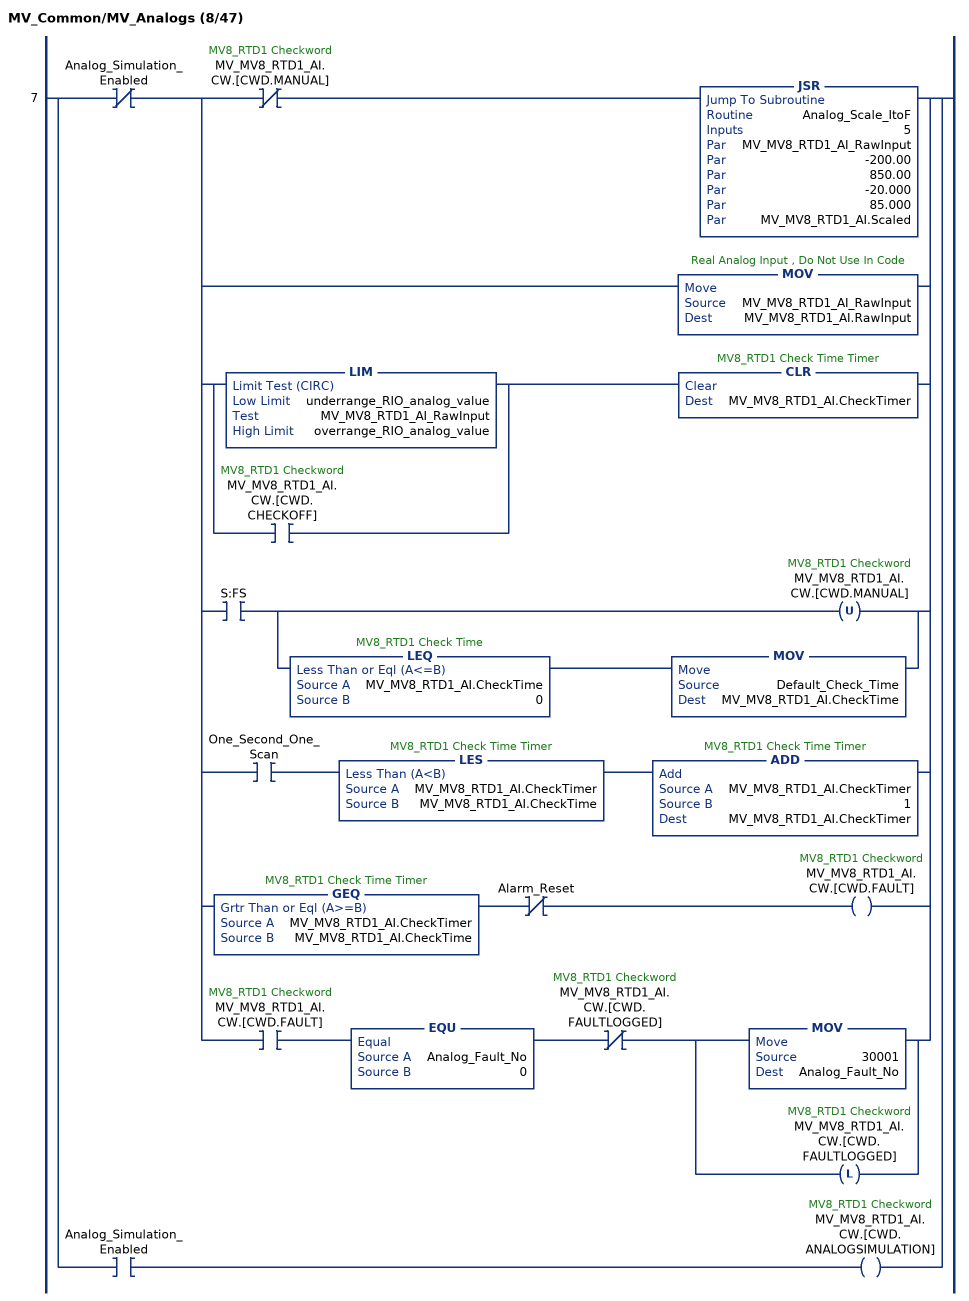
   7: [XIO(Analog_Simulation_Enabled) [XIO(MV_MV8_RTD1_AI.CW.[CWD.MANUAL]) JSR(Analog_Scale_ItoF,5,MV_MV8_RTD1_AI_RawInput,-200.00,850.00,-20.000,85.000,MV_MV8_RTD1_AI.Scaled) ,MOV(MV_MV8_RTD1_AI_RawInput,MV_MV8_RTD1_AI.RawInput) ,[LIM(underrange_RIO_analog_value,MV_MV8_RTD1_AI_RawInput,overrange_RIO_analog_value) ,XIC(MV_MV8_RTD1_AI.CW.[CWD.CHECKOFF]) ] CLR(MV_MV8_RTD1_AI.CheckTimer) ,XIC(S:FS) [OTU(MV_MV8_RTD1_AI.CW.[CWD.MANUAL]) ,LEQ(MV_MV8_RTD1_AI.CheckTime,0) MOV(Default_Check_Time,MV_MV8_RTD1_AI.CheckTime) ] ,XIC(One_Second_One_Scan) LES(MV_MV8_RTD1_AI.CheckTimer,MV_MV8_RTD1_AI.CheckTime) ADD(MV_MV8_RTD1_AI.CheckTimer,1,MV_MV8_RTD1_AI.CheckTimer) ,GEQ(MV_MV8_RTD1_AI.CheckTimer,MV_MV8_RTD1_AI.CheckTime) XIO(Alarm_Reset) OTE(MV_MV8_RTD1_AI.CW.[CWD.FAULT]) ,XIC(MV_MV8_RTD1_AI.CW.[CWD.FAULT]) EQU(Analog_Fault_No,0) XIO(MV_MV8_RTD1_AI.CW.[CWD.FAULTLOGGED]) [MOV(30001,Analog_Fault_No) ,OTL(MV_MV8_RTD1_AI.CW.[CWD.FAULTLOGGED]) ] ] ,XIC(Analog_Simulation_Enabled) OTE(MV_MV8_RTD1_AI.CW.[CWD.ANALOGSIMULATION]) ];
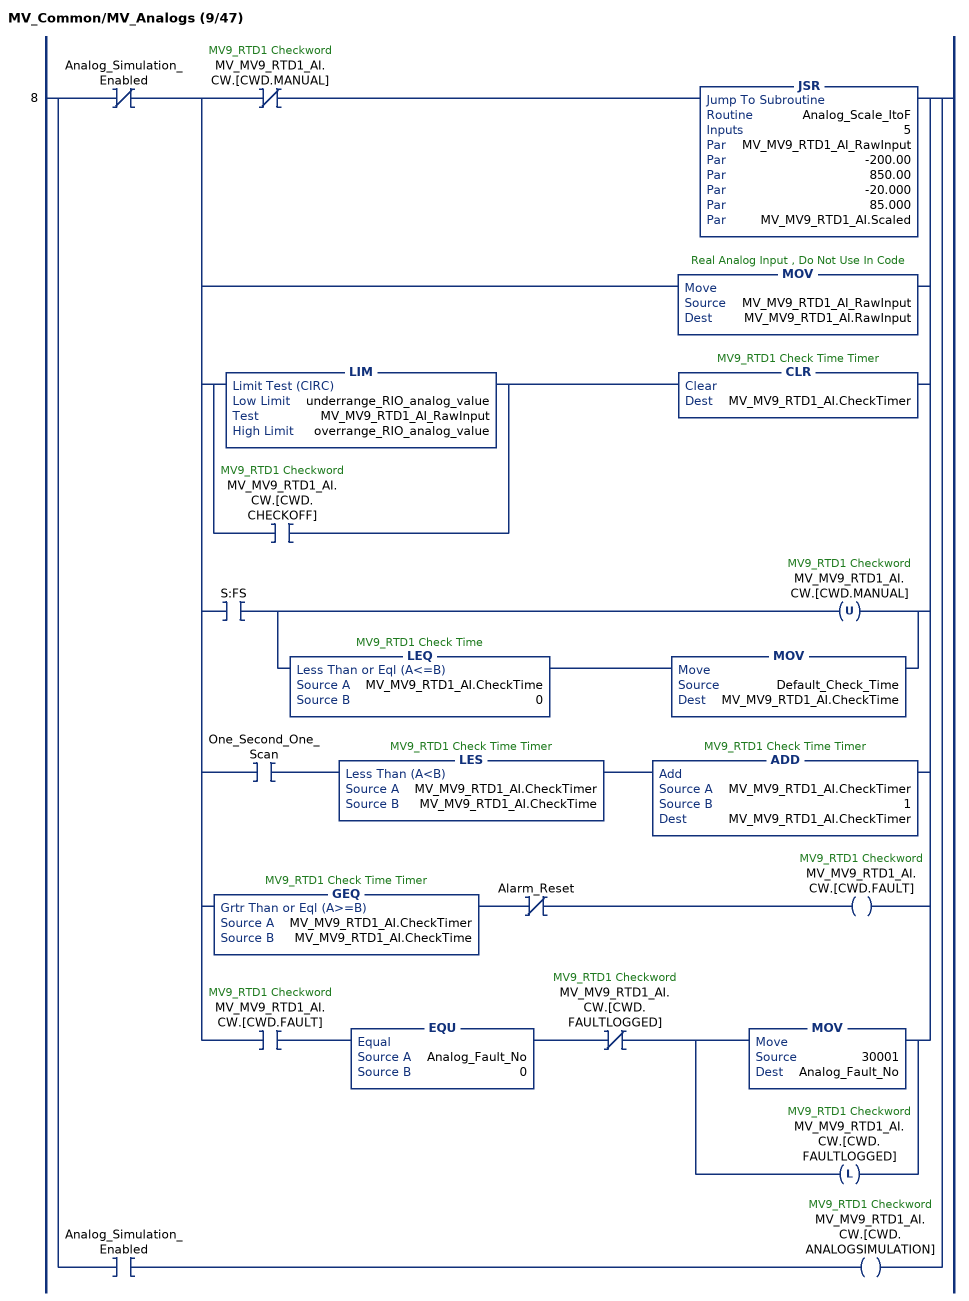
   8: [XIO(Analog_Simulation_Enabled) [XIO(MV_MV9_RTD1_AI.CW.[CWD.MANUAL]) JSR(Analog_Scale_ItoF,5,MV_MV9_RTD1_AI_RawInput,-200.00,850.00,-20.000,85.000,MV_MV9_RTD1_AI.Scaled) ,MOV(MV_MV9_RTD1_AI_RawInput,MV_MV9_RTD1_AI.RawInput) ,[LIM(underrange_RIO_analog_value,MV_MV9_RTD1_AI_RawInput,overrange_RIO_analog_value) ,XIC(MV_MV9_RTD1_AI.CW.[CWD.CHECKOFF]) ] CLR(MV_MV9_RTD1_AI.CheckTimer) ,XIC(S:FS) [OTU(MV_MV9_RTD1_AI.CW.[CWD.MANUAL]) ,LEQ(MV_MV9_RTD1_AI.CheckTime,0) MOV(Default_Check_Time,MV_MV9_RTD1_AI.CheckTime) ] ,XIC(One_Second_One_Scan) LES(MV_MV9_RTD1_AI.CheckTimer,MV_MV9_RTD1_AI.CheckTime) ADD(MV_MV9_RTD1_AI.CheckTimer,1,MV_MV9_RTD1_AI.CheckTimer) ,GEQ(MV_MV9_RTD1_AI.CheckTimer,MV_MV9_RTD1_AI.CheckTime) XIO(Alarm_Reset) OTE(MV_MV9_RTD1_AI.CW.[CWD.FAULT]) ,XIC(MV_MV9_RTD1_AI.CW.[CWD.FAULT]) EQU(Analog_Fault_No,0) XIO(MV_MV9_RTD1_AI.CW.[CWD.FAULTLOGGED]) [MOV(30001,Analog_Fault_No) ,OTL(MV_MV9_RTD1_AI.CW.[CWD.FAULTLOGGED]) ] ] ,XIC(Analog_Simulation_Enabled) OTE(MV_MV9_RTD1_AI.CW.[CWD.ANALOGSIMULATION]) ];
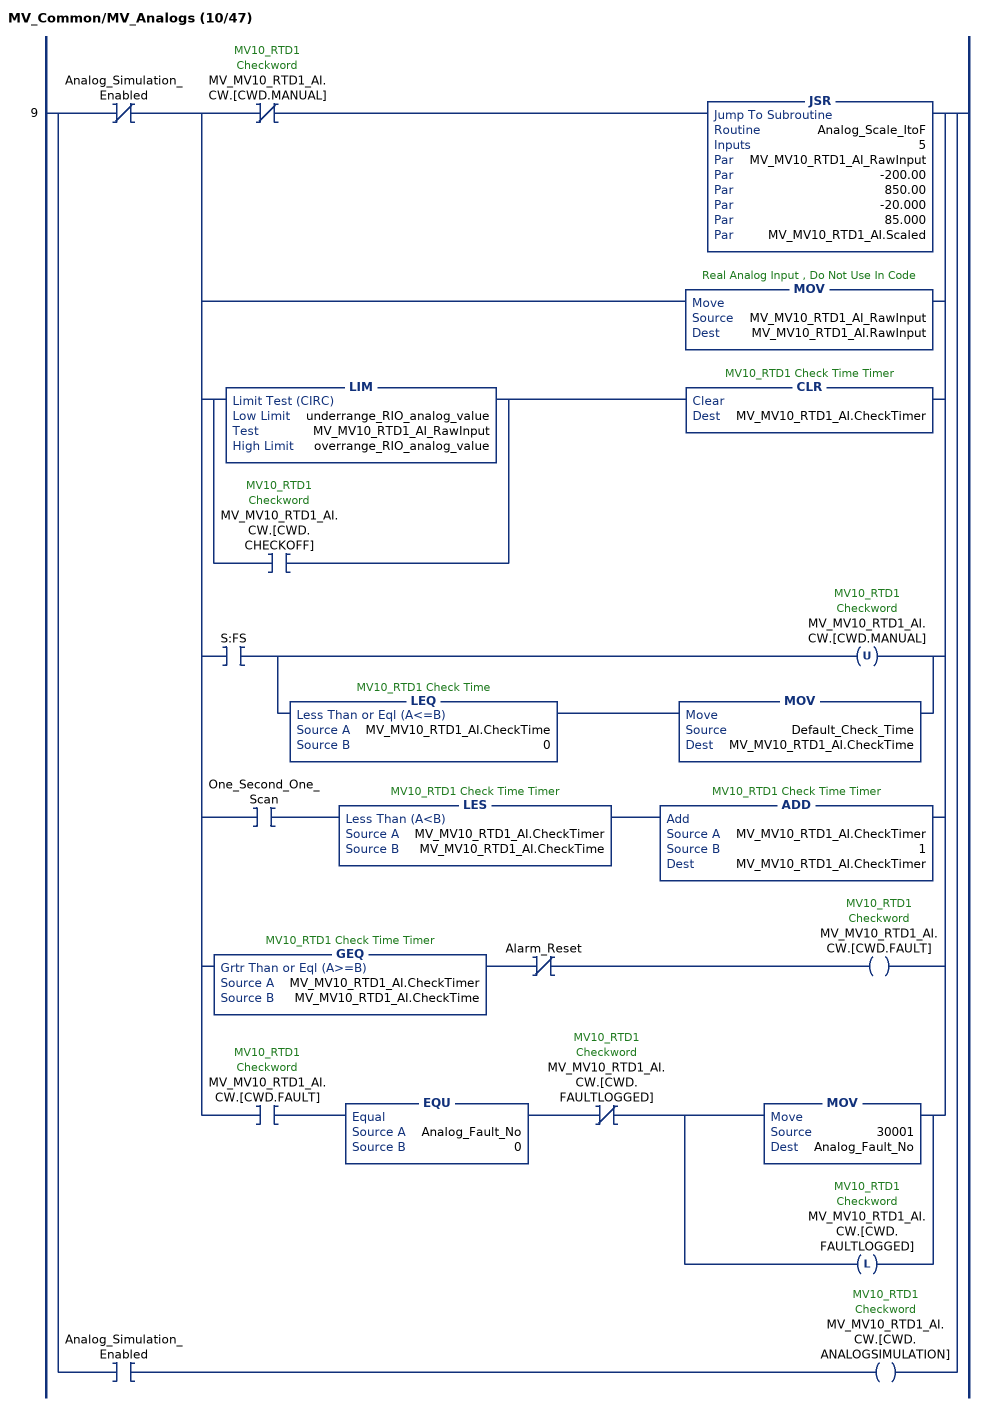
   9: [XIO(Analog_Simulation_Enabled) [XIO(MV_MV10_RTD1_AI.CW.[CWD.MANUAL]) JSR(Analog_Scale_ItoF,5,MV_MV10_RTD1_AI_RawInput,-200.00,850.00,-20.000,85.000,MV_MV10_RTD1_AI.Scaled) ,MOV(MV_MV10_RTD1_AI_RawInput,MV_MV10_RTD1_AI.RawInput) ,[LIM(underrange_RIO_analog_value,MV_MV10_RTD1_AI_RawInput,overrange_RIO_analog_value) ,XIC(MV_MV10_RTD1_AI.CW.[CWD.CHECKOFF]) ] CLR(MV_MV10_RTD1_AI.CheckTimer) ,XIC(S:FS) [OTU(MV_MV10_RTD1_AI.CW.[CWD.MANUAL]) ,LEQ(MV_MV10_RTD1_AI.CheckTime,0) MOV(Default_Check_Time,MV_MV10_RTD1_AI.CheckTime) ] ,XIC(One_Second_One_Scan) LES(MV_MV10_RTD1_AI.CheckTimer,MV_MV10_RTD1_AI.CheckTime) ADD(MV_MV10_RTD1_AI.CheckTimer,1,MV_MV10_RTD1_AI.CheckTimer) ,GEQ(MV_MV10_RTD1_AI.CheckTimer,MV_MV10_RTD1_AI.CheckTime) XIO(Alarm_Reset) OTE(MV_MV10_RTD1_AI.CW.[CWD.FAULT]) ,XIC(MV_MV10_RTD1_AI.CW.[CWD.FAULT]) EQU(Analog_Fault_No,0) XIO(MV_MV10_RTD1_AI.CW.[CWD.FAULTLOGGED]) [MOV(30001,Analog_Fault_No) ,OTL(MV_MV10_RTD1_AI.CW.[CWD.FAULTLOGGED]) ] ] ,XIC(Analog_Simulation_Enabled) OTE(MV_MV10_RTD1_AI.CW.[CWD.ANALOGSIMULATION]) ];
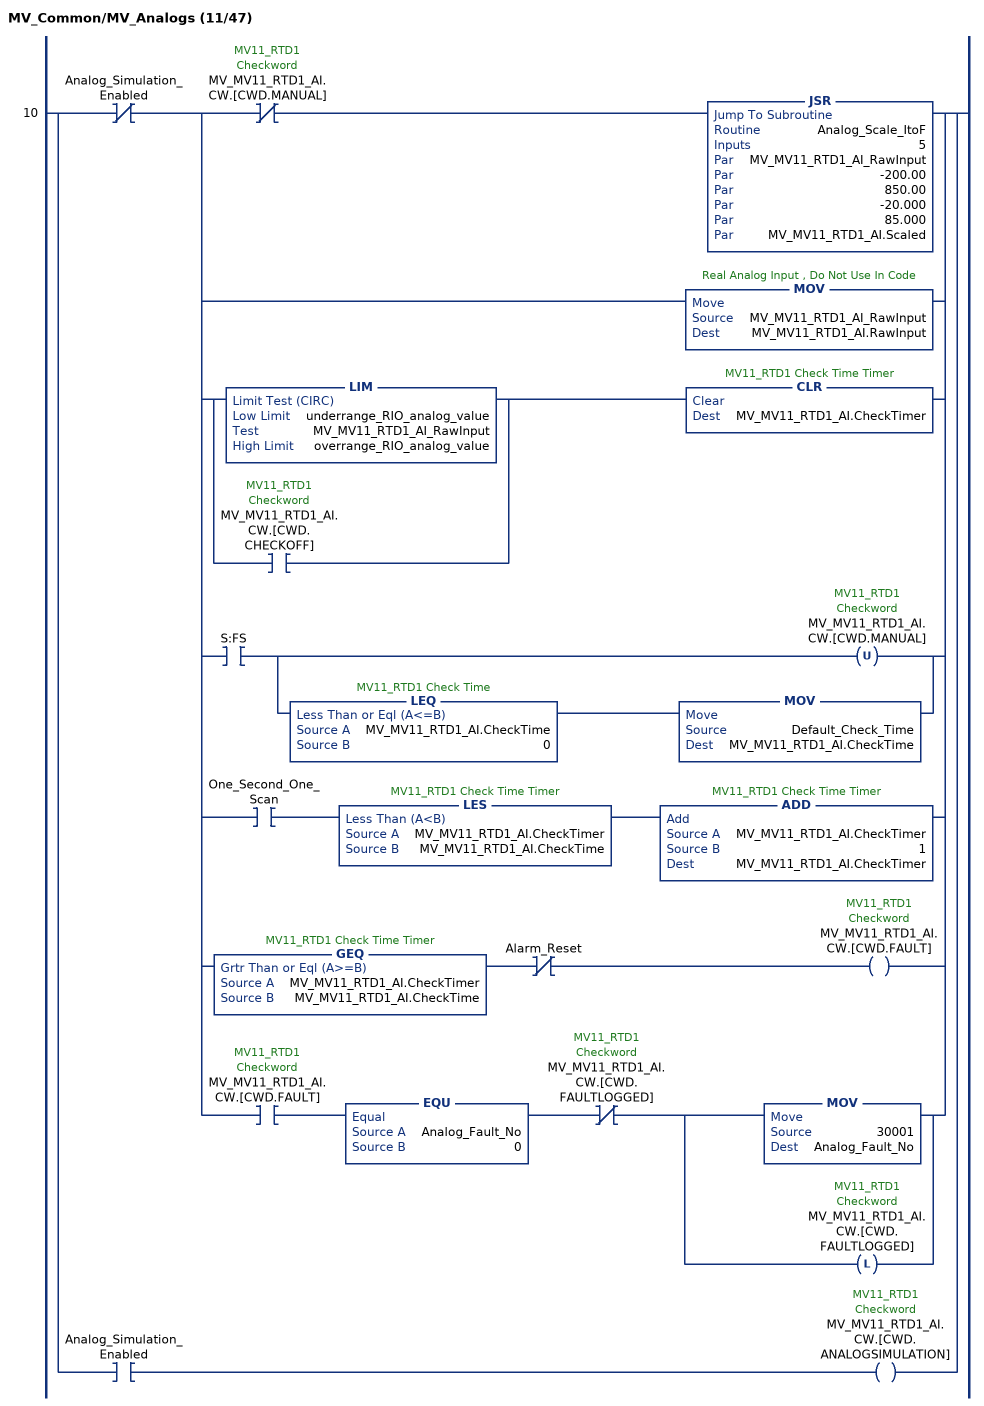
   10: [XIO(Analog_Simulation_Enabled) [XIO(MV_MV11_RTD1_AI.CW.[CWD.MANUAL]) JSR(Analog_Scale_ItoF,5,MV_MV11_RTD1_AI_RawInput,-200.00,850.00,-20.000,85.000,MV_MV11_RTD1_AI.Scaled) ,MOV(MV_MV11_RTD1_AI_RawInput,MV_MV11_RTD1_AI.RawInput) ,[LIM(underrange_RIO_analog_value,MV_MV11_RTD1_AI_RawInput,overrange_RIO_analog_value) ,XIC(MV_MV11_RTD1_AI.CW.[CWD.CHECKOFF]) ] CLR(MV_MV11_RTD1_AI.CheckTimer) ,XIC(S:FS) [OTU(MV_MV11_RTD1_AI.CW.[CWD.MANUAL]) ,LEQ(MV_MV11_RTD1_AI.CheckTime,0) MOV(Default_Check_Time,MV_MV11_RTD1_AI.CheckTime) ] ,XIC(One_Second_One_Scan) LES(MV_MV11_RTD1_AI.CheckTimer,MV_MV11_RTD1_AI.CheckTime) ADD(MV_MV11_RTD1_AI.CheckTimer,1,MV_MV11_RTD1_AI.CheckTimer) ,GEQ(MV_MV11_RTD1_AI.CheckTimer,MV_MV11_RTD1_AI.CheckTime) XIO(Alarm_Reset) OTE(MV_MV11_RTD1_AI.CW.[CWD.FAULT]) ,XIC(MV_MV11_RTD1_AI.CW.[CWD.FAULT]) EQU(Analog_Fault_No,0) XIO(MV_MV11_RTD1_AI.CW.[CWD.FAULTLOGGED]) [MOV(30001,Analog_Fault_No) ,OTL(MV_MV11_RTD1_AI.CW.[CWD.FAULTLOGGED]) ] ] ,XIC(Analog_Simulation_Enabled) OTE(MV_MV11_RTD1_AI.CW.[CWD.ANALOGSIMULATION]) ];
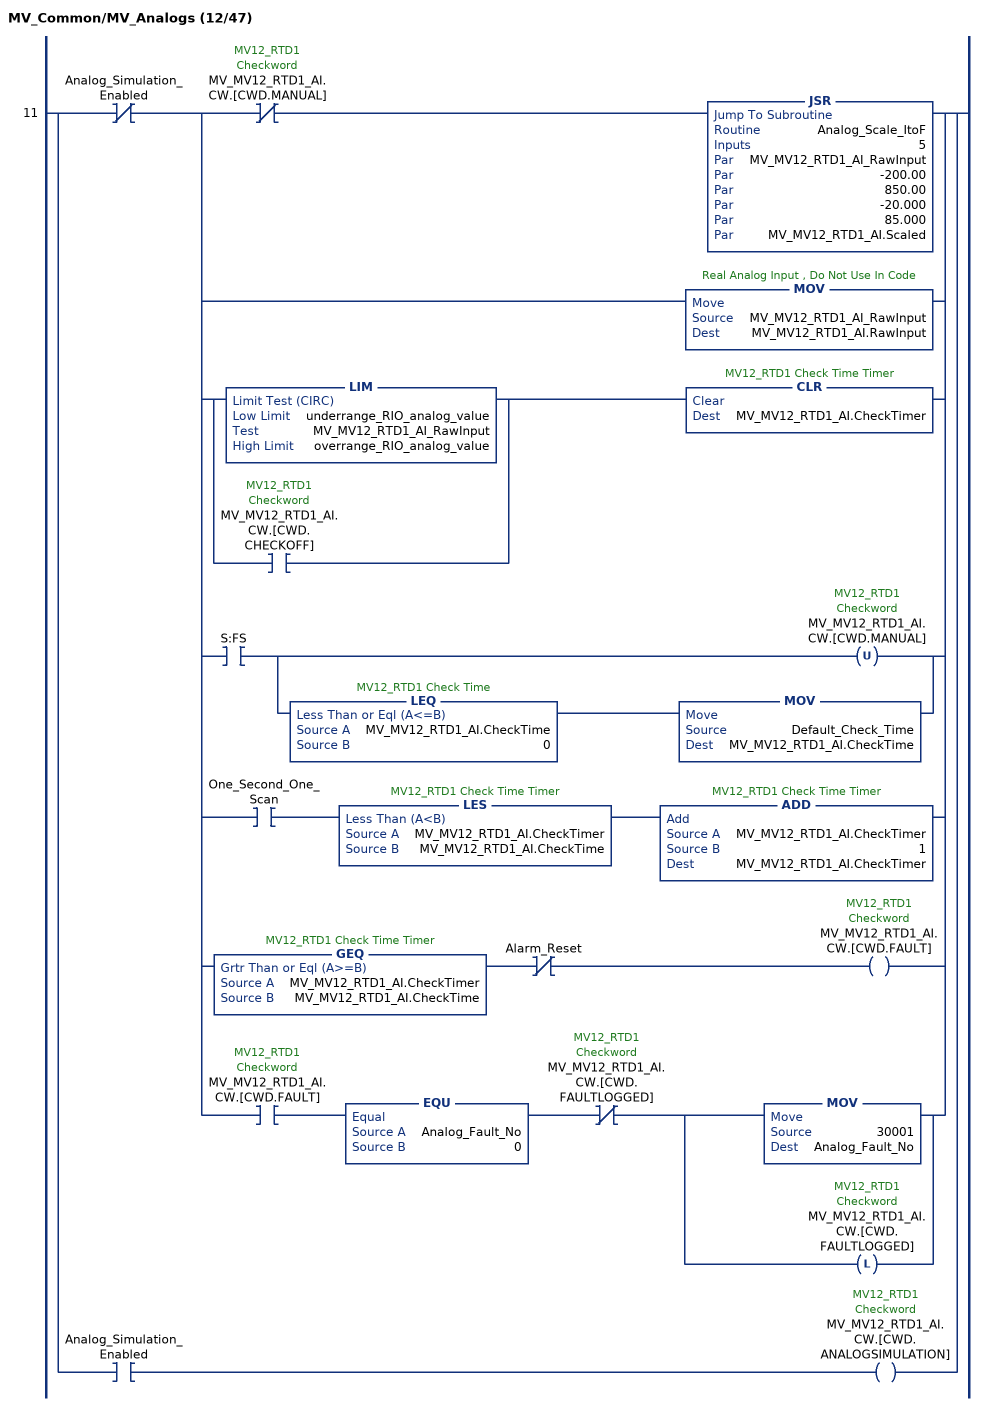
   11: [XIO(Analog_Simulation_Enabled) [XIO(MV_MV12_RTD1_AI.CW.[CWD.MANUAL]) JSR(Analog_Scale_ItoF,5,MV_MV12_RTD1_AI_RawInput,-200.00,850.00,-20.000,85.000,MV_MV12_RTD1_AI.Scaled) ,MOV(MV_MV12_RTD1_AI_RawInput,MV_MV12_RTD1_AI.RawInput) ,[LIM(underrange_RIO_analog_value,MV_MV12_RTD1_AI_RawInput,overrange_RIO_analog_value) ,XIC(MV_MV12_RTD1_AI.CW.[CWD.CHECKOFF]) ] CLR(MV_MV12_RTD1_AI.CheckTimer) ,XIC(S:FS) [OTU(MV_MV12_RTD1_AI.CW.[CWD.MANUAL]) ,LEQ(MV_MV12_RTD1_AI.CheckTime,0) MOV(Default_Check_Time,MV_MV12_RTD1_AI.CheckTime) ] ,XIC(One_Second_One_Scan) LES(MV_MV12_RTD1_AI.CheckTimer,MV_MV12_RTD1_AI.CheckTime) ADD(MV_MV12_RTD1_AI.CheckTimer,1,MV_MV12_RTD1_AI.CheckTimer) ,GEQ(MV_MV12_RTD1_AI.CheckTimer,MV_MV12_RTD1_AI.CheckTime) XIO(Alarm_Reset) OTE(MV_MV12_RTD1_AI.CW.[CWD.FAULT]) ,XIC(MV_MV12_RTD1_AI.CW.[CWD.FAULT]) EQU(Analog_Fault_No,0) XIO(MV_MV12_RTD1_AI.CW.[CWD.FAULTLOGGED]) [MOV(30001,Analog_Fault_No) ,OTL(MV_MV12_RTD1_AI.CW.[CWD.FAULTLOGGED]) ] ] ,XIC(Analog_Simulation_Enabled) OTE(MV_MV12_RTD1_AI.CW.[CWD.ANALOGSIMULATION]) ];
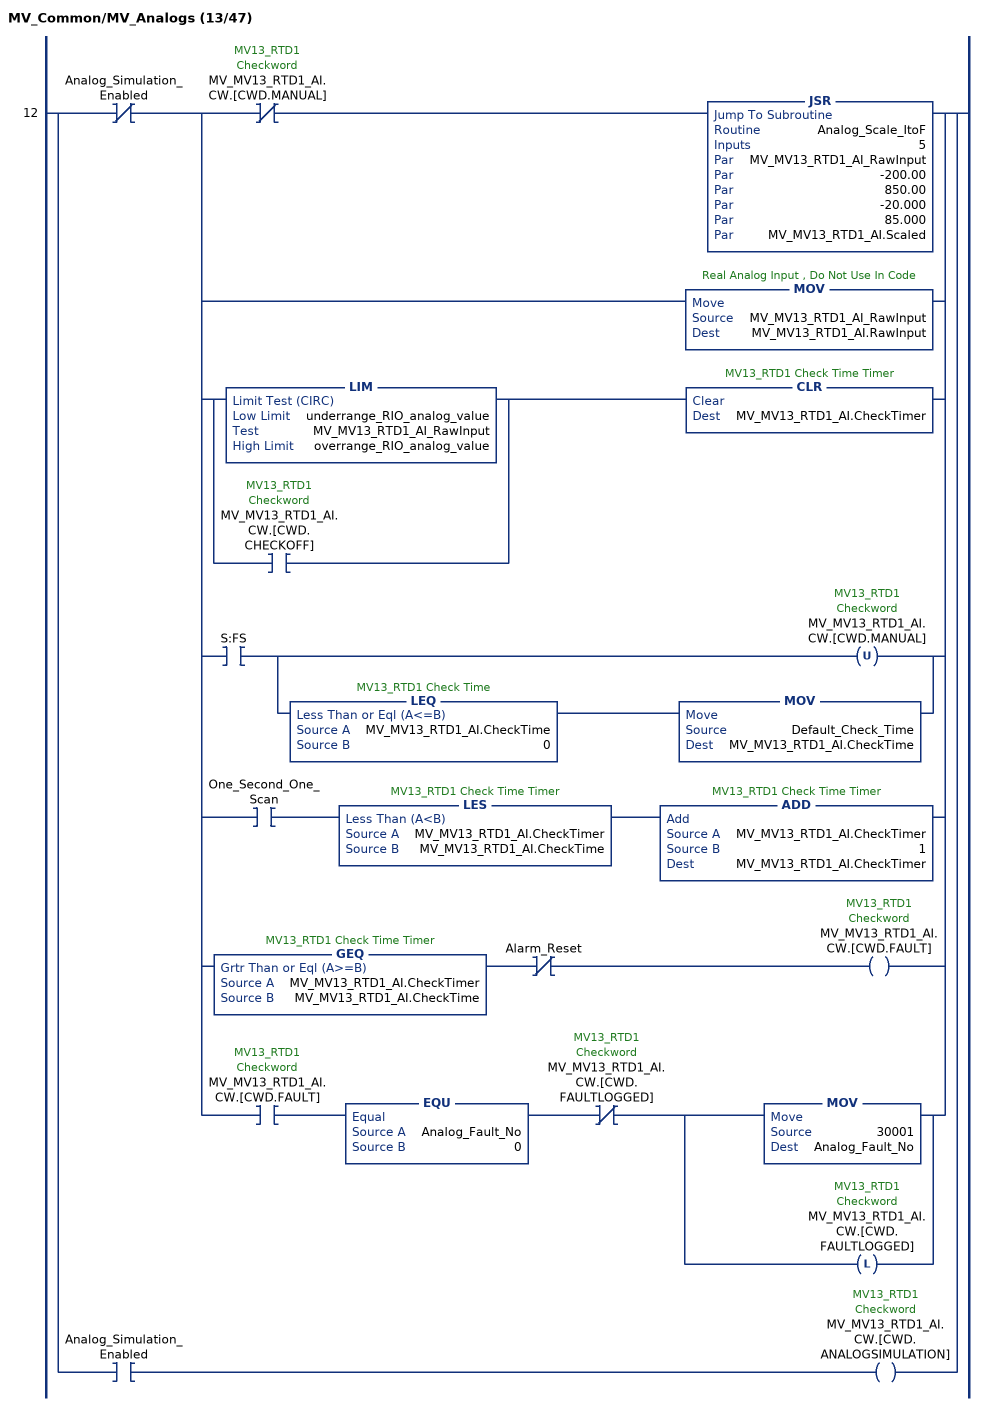
   12: [XIO(Analog_Simulation_Enabled) [XIO(MV_MV13_RTD1_AI.CW.[CWD.MANUAL]) JSR(Analog_Scale_ItoF,5,MV_MV13_RTD1_AI_RawInput,-200.00,850.00,-20.000,85.000,MV_MV13_RTD1_AI.Scaled) ,MOV(MV_MV13_RTD1_AI_RawInput,MV_MV13_RTD1_AI.RawInput) ,[LIM(underrange_RIO_analog_value,MV_MV13_RTD1_AI_RawInput,overrange_RIO_analog_value) ,XIC(MV_MV13_RTD1_AI.CW.[CWD.CHECKOFF]) ] CLR(MV_MV13_RTD1_AI.CheckTimer) ,XIC(S:FS) [OTU(MV_MV13_RTD1_AI.CW.[CWD.MANUAL]) ,LEQ(MV_MV13_RTD1_AI.CheckTime,0) MOV(Default_Check_Time,MV_MV13_RTD1_AI.CheckTime) ] ,XIC(One_Second_One_Scan) LES(MV_MV13_RTD1_AI.CheckTimer,MV_MV13_RTD1_AI.CheckTime) ADD(MV_MV13_RTD1_AI.CheckTimer,1,MV_MV13_RTD1_AI.CheckTimer) ,GEQ(MV_MV13_RTD1_AI.CheckTimer,MV_MV13_RTD1_AI.CheckTime) XIO(Alarm_Reset) OTE(MV_MV13_RTD1_AI.CW.[CWD.FAULT]) ,XIC(MV_MV13_RTD1_AI.CW.[CWD.FAULT]) EQU(Analog_Fault_No,0) XIO(MV_MV13_RTD1_AI.CW.[CWD.FAULTLOGGED]) [MOV(30001,Analog_Fault_No) ,OTL(MV_MV13_RTD1_AI.CW.[CWD.FAULTLOGGED]) ] ] ,XIC(Analog_Simulation_Enabled) OTE(MV_MV13_RTD1_AI.CW.[CWD.ANALOGSIMULATION]) ];
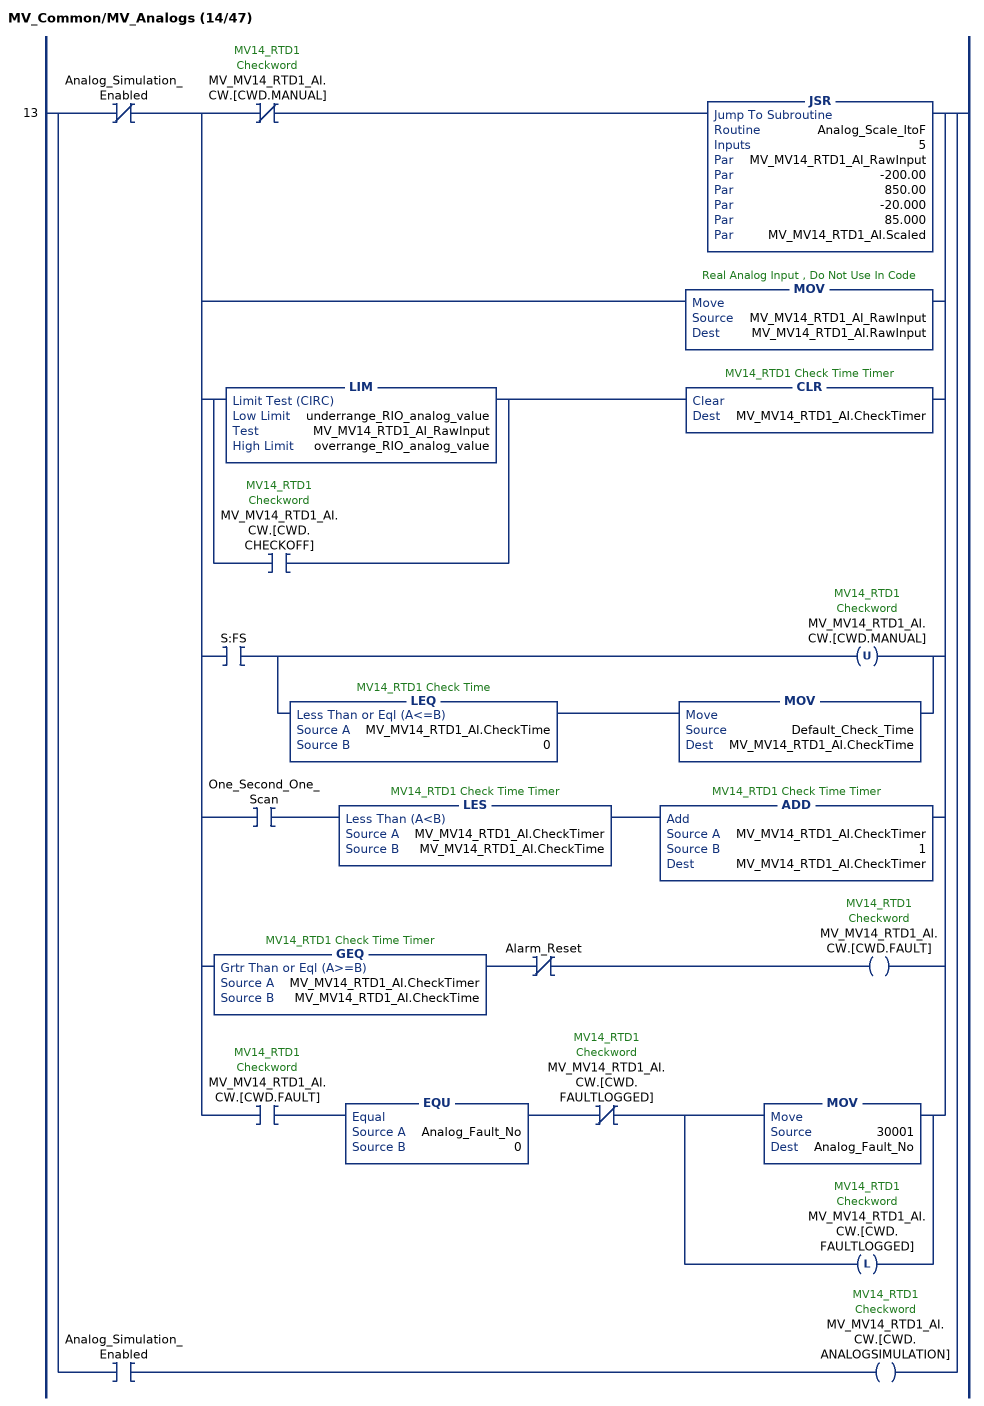
   13: [XIO(Analog_Simulation_Enabled) [XIO(MV_MV14_RTD1_AI.CW.[CWD.MANUAL]) JSR(Analog_Scale_ItoF,5,MV_MV14_RTD1_AI_RawInput,-200.00,850.00,-20.000,85.000,MV_MV14_RTD1_AI.Scaled) ,MOV(MV_MV14_RTD1_AI_RawInput,MV_MV14_RTD1_AI.RawInput) ,[LIM(underrange_RIO_analog_value,MV_MV14_RTD1_AI_RawInput,overrange_RIO_analog_value) ,XIC(MV_MV14_RTD1_AI.CW.[CWD.CHECKOFF]) ] CLR(MV_MV14_RTD1_AI.CheckTimer) ,XIC(S:FS) [OTU(MV_MV14_RTD1_AI.CW.[CWD.MANUAL]) ,LEQ(MV_MV14_RTD1_AI.CheckTime,0) MOV(Default_Check_Time,MV_MV14_RTD1_AI.CheckTime) ] ,XIC(One_Second_One_Scan) LES(MV_MV14_RTD1_AI.CheckTimer,MV_MV14_RTD1_AI.CheckTime) ADD(MV_MV14_RTD1_AI.CheckTimer,1,MV_MV14_RTD1_AI.CheckTimer) ,GEQ(MV_MV14_RTD1_AI.CheckTimer,MV_MV14_RTD1_AI.CheckTime) XIO(Alarm_Reset) OTE(MV_MV14_RTD1_AI.CW.[CWD.FAULT]) ,XIC(MV_MV14_RTD1_AI.CW.[CWD.FAULT]) EQU(Analog_Fault_No,0) XIO(MV_MV14_RTD1_AI.CW.[CWD.FAULTLOGGED]) [MOV(30001,Analog_Fault_No) ,OTL(MV_MV14_RTD1_AI.CW.[CWD.FAULTLOGGED]) ] ] ,XIC(Analog_Simulation_Enabled) OTE(MV_MV14_RTD1_AI.CW.[CWD.ANALOGSIMULATION]) ];
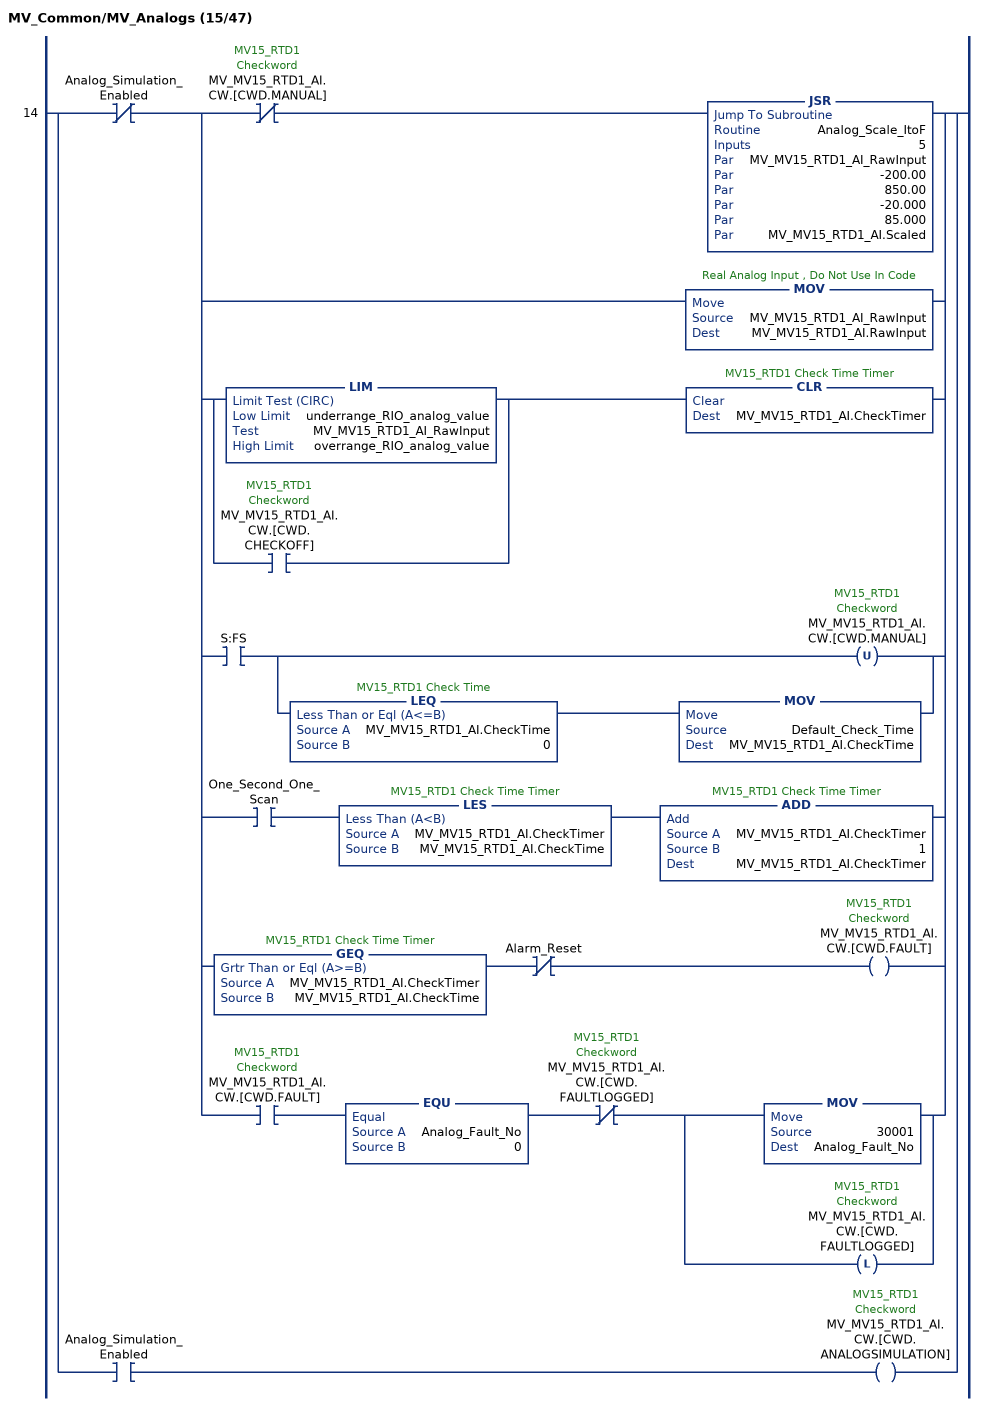
   14: [XIO(Analog_Simulation_Enabled) [XIO(MV_MV15_RTD1_AI.CW.[CWD.MANUAL]) JSR(Analog_Scale_ItoF,5,MV_MV15_RTD1_AI_RawInput,-200.00,850.00,-20.000,85.000,MV_MV15_RTD1_AI.Scaled) ,MOV(MV_MV15_RTD1_AI_RawInput,MV_MV15_RTD1_AI.RawInput) ,[LIM(underrange_RIO_analog_value,MV_MV15_RTD1_AI_RawInput,overrange_RIO_analog_value) ,XIC(MV_MV15_RTD1_AI.CW.[CWD.CHECKOFF]) ] CLR(MV_MV15_RTD1_AI.CheckTimer) ,XIC(S:FS) [OTU(MV_MV15_RTD1_AI.CW.[CWD.MANUAL]) ,LEQ(MV_MV15_RTD1_AI.CheckTime,0) MOV(Default_Check_Time,MV_MV15_RTD1_AI.CheckTime) ] ,XIC(One_Second_One_Scan) LES(MV_MV15_RTD1_AI.CheckTimer,MV_MV15_RTD1_AI.CheckTime) ADD(MV_MV15_RTD1_AI.CheckTimer,1,MV_MV15_RTD1_AI.CheckTimer) ,GEQ(MV_MV15_RTD1_AI.CheckTimer,MV_MV15_RTD1_AI.CheckTime) XIO(Alarm_Reset) OTE(MV_MV15_RTD1_AI.CW.[CWD.FAULT]) ,XIC(MV_MV15_RTD1_AI.CW.[CWD.FAULT]) EQU(Analog_Fault_No,0) XIO(MV_MV15_RTD1_AI.CW.[CWD.FAULTLOGGED]) [MOV(30001,Analog_Fault_No) ,OTL(MV_MV15_RTD1_AI.CW.[CWD.FAULTLOGGED]) ] ] ,XIC(Analog_Simulation_Enabled) OTE(MV_MV15_RTD1_AI.CW.[CWD.ANALOGSIMULATION]) ];
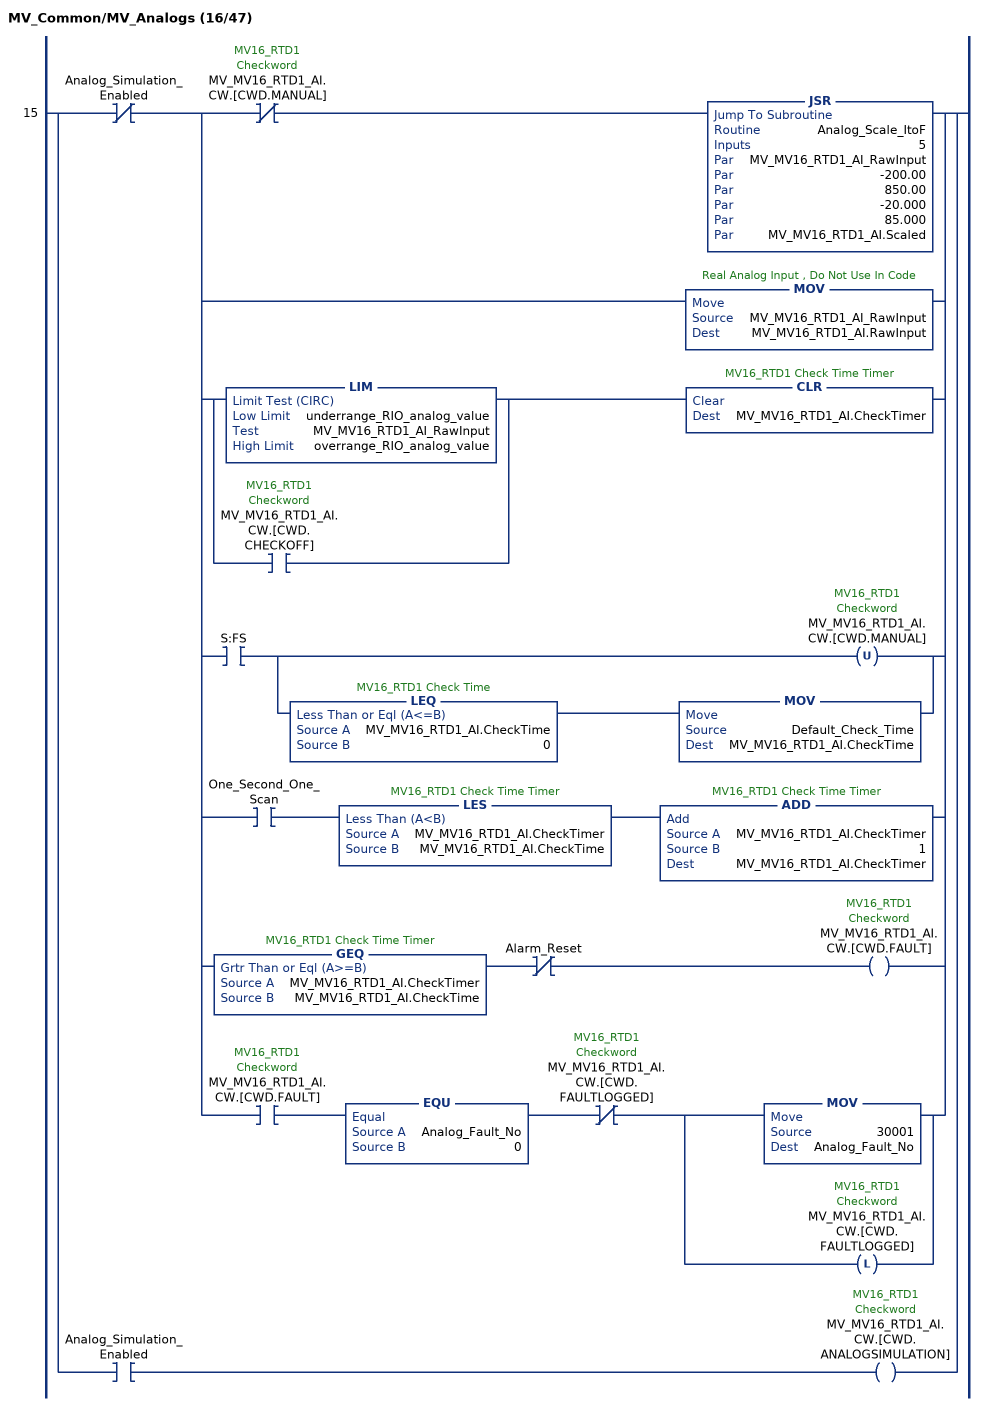
   15: [XIO(Analog_Simulation_Enabled) [XIO(MV_MV16_RTD1_AI.CW.[CWD.MANUAL]) JSR(Analog_Scale_ItoF,5,MV_MV16_RTD1_AI_RawInput,-200.00,850.00,-20.000,85.000,MV_MV16_RTD1_AI.Scaled) ,MOV(MV_MV16_RTD1_AI_RawInput,MV_MV16_RTD1_AI.RawInput) ,[LIM(underrange_RIO_analog_value,MV_MV16_RTD1_AI_RawInput,overrange_RIO_analog_value) ,XIC(MV_MV16_RTD1_AI.CW.[CWD.CHECKOFF]) ] CLR(MV_MV16_RTD1_AI.CheckTimer) ,XIC(S:FS) [OTU(MV_MV16_RTD1_AI.CW.[CWD.MANUAL]) ,LEQ(MV_MV16_RTD1_AI.CheckTime,0) MOV(Default_Check_Time,MV_MV16_RTD1_AI.CheckTime) ] ,XIC(One_Second_One_Scan) LES(MV_MV16_RTD1_AI.CheckTimer,MV_MV16_RTD1_AI.CheckTime) ADD(MV_MV16_RTD1_AI.CheckTimer,1,MV_MV16_RTD1_AI.CheckTimer) ,GEQ(MV_MV16_RTD1_AI.CheckTimer,MV_MV16_RTD1_AI.CheckTime) XIO(Alarm_Reset) OTE(MV_MV16_RTD1_AI.CW.[CWD.FAULT]) ,XIC(MV_MV16_RTD1_AI.CW.[CWD.FAULT]) EQU(Analog_Fault_No,0) XIO(MV_MV16_RTD1_AI.CW.[CWD.FAULTLOGGED]) [MOV(30001,Analog_Fault_No) ,OTL(MV_MV16_RTD1_AI.CW.[CWD.FAULTLOGGED]) ] ] ,XIC(Analog_Simulation_Enabled) OTE(MV_MV16_RTD1_AI.CW.[CWD.ANALOGSIMULATION]) ];
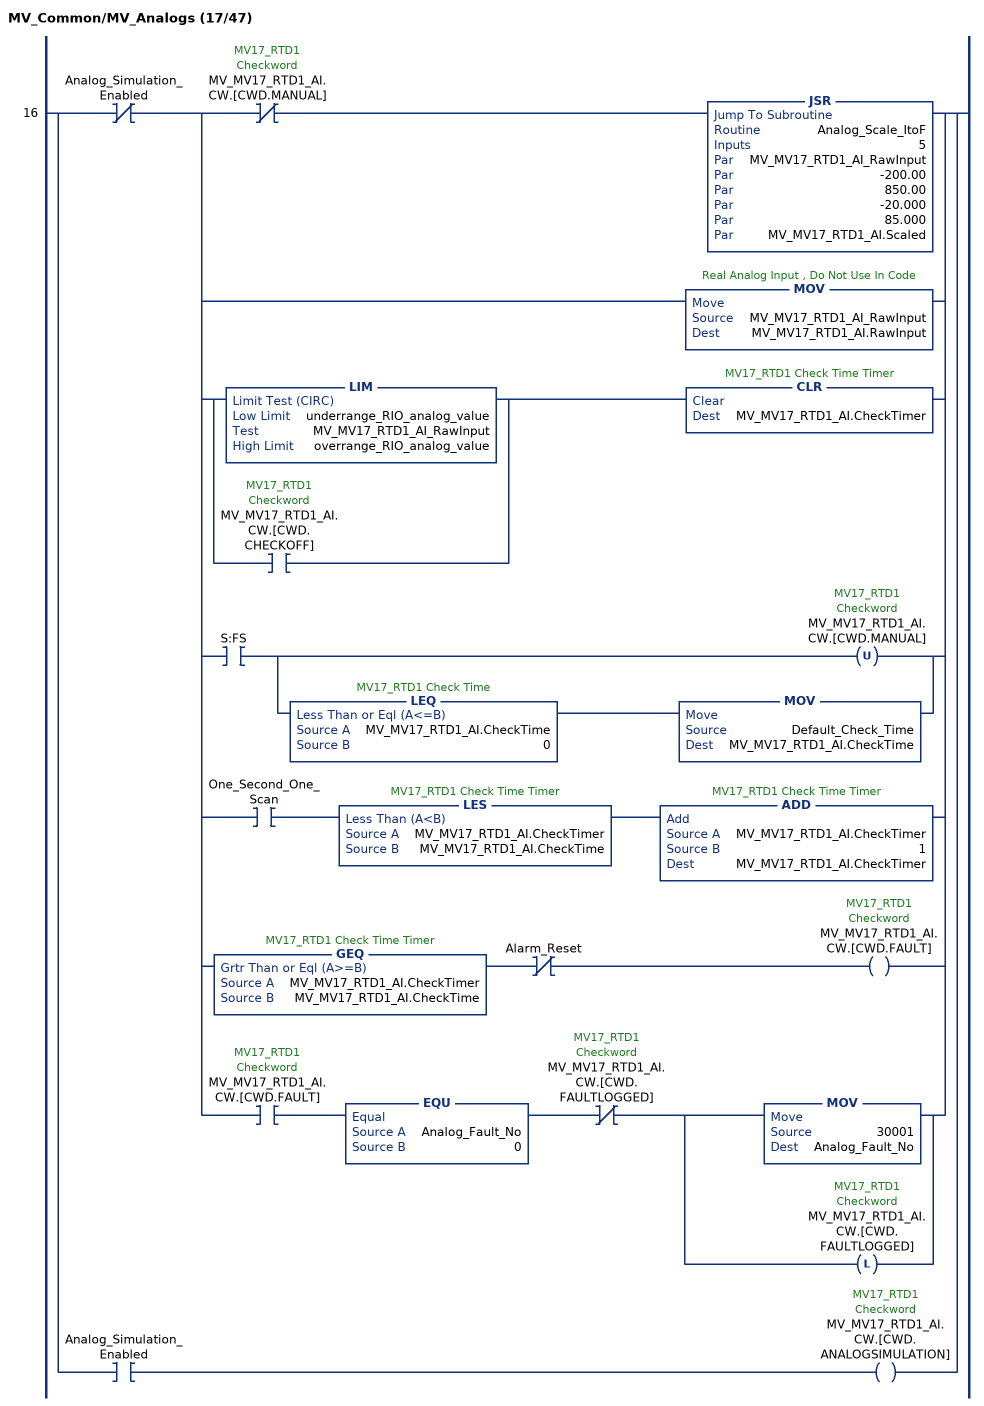
   16: [XIO(Analog_Simulation_Enabled) [XIO(MV_MV17_RTD1_AI.CW.[CWD.MANUAL]) JSR(Analog_Scale_ItoF,5,MV_MV17_RTD1_AI_RawInput,-200.00,850.00,-20.000,85.000,MV_MV17_RTD1_AI.Scaled) ,MOV(MV_MV17_RTD1_AI_RawInput,MV_MV17_RTD1_AI.RawInput) ,[LIM(underrange_RIO_analog_value,MV_MV17_RTD1_AI_RawInput,overrange_RIO_analog_value) ,XIC(MV_MV17_RTD1_AI.CW.[CWD.CHECKOFF]) ] CLR(MV_MV17_RTD1_AI.CheckTimer) ,XIC(S:FS) [OTU(MV_MV17_RTD1_AI.CW.[CWD.MANUAL]) ,LEQ(MV_MV17_RTD1_AI.CheckTime,0) MOV(Default_Check_Time,MV_MV17_RTD1_AI.CheckTime) ] ,XIC(One_Second_One_Scan) LES(MV_MV17_RTD1_AI.CheckTimer,MV_MV17_RTD1_AI.CheckTime) ADD(MV_MV17_RTD1_AI.CheckTimer,1,MV_MV17_RTD1_AI.CheckTimer) ,GEQ(MV_MV17_RTD1_AI.CheckTimer,MV_MV17_RTD1_AI.CheckTime) XIO(Alarm_Reset) OTE(MV_MV17_RTD1_AI.CW.[CWD.FAULT]) ,XIC(MV_MV17_RTD1_AI.CW.[CWD.FAULT]) EQU(Analog_Fault_No,0) XIO(MV_MV17_RTD1_AI.CW.[CWD.FAULTLOGGED]) [MOV(30001,Analog_Fault_No) ,OTL(MV_MV17_RTD1_AI.CW.[CWD.FAULTLOGGED]) ] ] ,XIC(Analog_Simulation_Enabled) OTE(MV_MV17_RTD1_AI.CW.[CWD.ANALOGSIMULATION]) ];
